// TIA Portal project "Inteligenta_szklarnia" (V15.1)

(* hardware
DEVICE "HMI_test"  KTP700 Basic PN
   slot 0: "HMI_test"  KTP700 Basic PN  6AV2 123-2GB03-0AX0  15.1.0.0
   slot 1: "HMI_RT_1"  KTP700 Basic PN  6AV2 123-2GB03-0AX0  15.1.0.0
   slot 5: "HMI_test.IE_CP_1"  PROFINET Interface  15.0.1.0
      slot 1: "PROFINET Interface_1"  PROFINET Interface
         slot 1: "Port_1"  Port
DEVICE "S7-1200 station_2"  S7-1200 Station
   slot 0: "Rack_0"  S7-1200 Rack  Rack  V1.0
   slot 1: "PLC_1"  CPU 1214C AC/DC/Rly  6ES7 214-1BE30-0XB0  V2.2
DEVICE "HMI_1"  KTP700 Basic PN
   slot 0: "HMI_1"  KTP700 Basic PN  6AV2 123-2GB03-0AX0  15.1.0.0
   slot 1: "HMI_RT_3"  KTP700 Basic PN  6AV2 123-2GB03-0AX0  15.1.0.0
   slot 5: "HMI_1.IE_CP_1"  PROFINET Interface  15.0.1.0
      slot 1: "PROFINET Interface_1"  PROFINET Interface
         slot 1: "Port_1"  Port
DEVICE "S7-1200 station_1"  S7-1200 Station
   slot 0: "Rack_0"  S7-1200 Rack  Rack  V1.0
   slot 1: "PLC_do_symulacji"  CPU 1214C AC/DC/Rly  6ES7 214-1BG40-0XB0  V4.2
DEVICE "HMI_do_symulacji"  KTP700 Basic PN
   slot 0: "HMI_do_symulacji"  KTP700 Basic PN  6AV2 123-2GB03-0AX0  15.1.0.0
   slot 1: "HMI_RT_2"  KTP700 Basic PN  6AV2 123-2GB03-0AX0  15.1.0.0
   slot 5: "HMI_do_symulacji.IE_CP_1"  PROFINET Interface  15.0.1.0
      slot 1: "PROFINET Interface_1"  PROFINET Interface
         slot 1: "Port_1"  Port
*)

// ===== PLC "PLC_1"  CPU 1214C AC/DC/Rly =====

VAR_GLOBAL   // PLC tag table "Default tag table"
   "Tag_1" AT %I0.0 : Bool;
   "Tag_ScreenNumber" AT %MD0 : DInt;
   "FirstScan" AT %M1.0 : Bool;
   "DiagStatusUpdate" AT %M1.1 : Bool;
   "AlwaysTRUE" AT %M1.2 : Bool;
   "AlwaysFALSE" AT %M1.3 : Bool;
END_VAR

VAR_GLOBAL   // PLC tag table "wyjscia"
   "Grzałka" AT %Q0.0 : Bool;
   "Wentylator" AT %Q0.1 : Bool;
   "Pompa_wodna" AT %Q0.2 : Bool;
   "Rolety_zamykanie" AT %Q0.4 : Bool;
   "Alarm_ostrzegwaczy" AT %Q0.5 : Bool;
   "Siłownik_okien_otwieranie" AT %Q0.6 : Bool;
   "Siłownik_okien_zamykanie" AT %Q0.7 : Bool;
   "Rolety_otwieranie" AT %Q0.3 : Bool;
END_VAR

DATA_BLOCK "Parametry"   // DB1
{ S7_Optimized_Access := 'TRUE' }
VERSION : 0.1
   VAR
      Wilgotność_powietrza : Int;
      Wilgotność_gleby : Int;
      temeratura : Real;
      Czujnik_światła : Int;
      Czujnik_wiatru : Int;
      czujnik_CO2 : Int;
      stopien_zasloniecia_rolet : Int;
   END_VAR
BEGIN
END_DATA_BLOCK

DATA_BLOCK "Wejscia_HMI"   // DB2
{ S7_Optimized_Access := 'TRUE' }
VERSION : 0.1
   VAR
      Temperatura : Real;
      CO2 : Real;
      Wilgotność_gleby : Int;
      Wilgotność_powietrza : Int;
      Zaciemnienie : Int;
      naslonecznienie_manual : Int;
   END_VAR
BEGIN
END_DATA_BLOCK

DATA_BLOCK "Receptury"   // DB3
{ S7_Optimized_Access := 'TRUE' }
VERSION : 0.1
   VAR
      nasłonecznienie : Array[0..5] of Int;
      system_okien : Array[0..5] of Bool;
      wilgotnosc_gleby : Array[0..5] of Int;
      wilgotnosc_powietrza : Array[0..5] of Int;
      temperatua : Array[0..5] of Real;
      nazwa : Array[0..5] of String;
   END_VAR
BEGIN
END_DATA_BLOCK

DATA_BLOCK "Archiwizowane_parametry"   // DB4
{ S7_Optimized_Access := 'TRUE' }
VERSION : 0.1
   VAR
      Temperatura : Array[0..335] of Real;
      Wilgotnosc : Array[0..335] of Int;
      Naslonecznienie : Array[0..335] of Int;
      iterator : Int := 0;   // Iterator służący do zapisu danych w odpowiednich komórkach tablicy.
      Zerowanie : Array[0..335] of Int;
   END_VAR
BEGIN
   Naslonecznienie[0] := 0;
   Naslonecznienie[1] := 0;
END_DATA_BLOCK

// folder: System blocks/Program resources

DATA_BLOCK "IEC_Timer_0_DB"   // DB5
{ S7_Optimized_Access := 'TRUE' }
AUTHOR : Simatic
FAMILY : IEC
NAME : IEC_TMR
VERSION : 1.0
// stored: InstanceOfName IEC_TIMER
"IEC_TIMER"
BEGIN
END_DATA_BLOCK

// folder: (top level)

FUNCTION "Rolety" : Void   // FC1, LAD
{ S7_Optimized_Access := 'TRUE' }
VERSION : 0.1
   VAR_INPUT
      Czy_automatyczny : Bool;
      Czy_manualny : Bool;
   END_VAR
   VAR_TEMP   // added for the SCL form of the ladder/FBD networks
      _w1 : Bool;
   END_VAR
BEGIN

REGION Network 1: Sterowanie roletami w trybie automatycznym
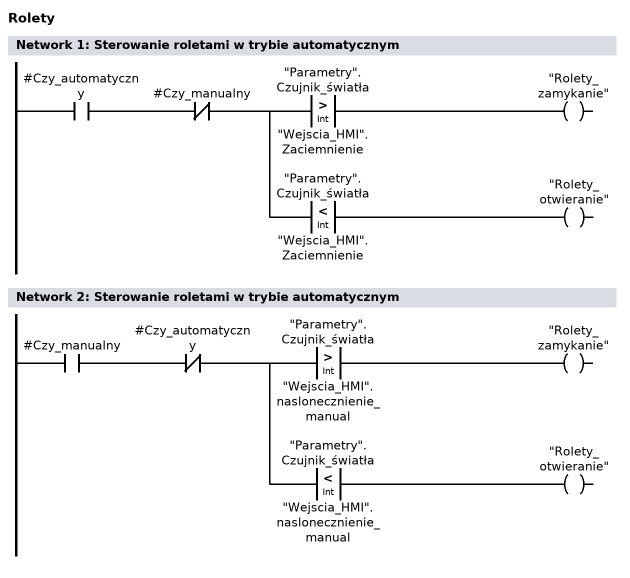
   RUNG wire#powerrail
      Contact( #Czy_automatyczny )
      I_Contact( #Czy_manualny )
      wire#w1
      { S7_Templates := "SrcType := Int" } GT_Contact(in1 := "Parametry".Czujnik_światła, in2 := "Wejscia_HMI".Zaciemnienie)
      Coil( "Rolety_zamykanie" )
   END_RUNG
   RUNG wire#w1
      { S7_Templates := "SrcType := Int" } LT_Contact(in1 := "Parametry".Czujnik_światła, in2 := "Wejscia_HMI".Zaciemnienie)
      Coil( "Rolety_otwieranie" )
   END_RUNG
   // the same network as SCL:
   #_w1 := #Czy_automatyczny AND NOT #Czy_manualny;
   "Rolety_zamykanie" := #_w1 AND ("Parametry".Czujnik_światła > "Wejscia_HMI".Zaciemnienie);
   "Rolety_otwieranie" := #_w1 AND ("Parametry".Czujnik_światła < "Wejscia_HMI".Zaciemnienie);
END_REGION

REGION Network 2: Sterowanie roletami w trybie automatycznym
   RUNG wire#powerrail
      Contact( #Czy_manualny )
      I_Contact( #Czy_automatyczny )
      wire#w1
      { S7_Templates := "SrcType := Int" } GT_Contact(in1 := "Parametry".Czujnik_światła, in2 := "Wejscia_HMI".naslonecznienie_manual)
      Coil( "Rolety_zamykanie" )
   END_RUNG
   RUNG wire#w1
      { S7_Templates := "SrcType := Int" } LT_Contact(in1 := "Parametry".Czujnik_światła, in2 := "Wejscia_HMI".naslonecznienie_manual)
      Coil( "Rolety_otwieranie" )
   END_RUNG
   // the same network as SCL:
   #_w1 := #Czy_manualny AND NOT #Czy_automatyczny;
   "Rolety_zamykanie" := #_w1 AND ("Parametry".Czujnik_światła > "Wejscia_HMI".naslonecznienie_manual);
   "Rolety_otwieranie" := #_w1 AND ("Parametry".Czujnik_światła < "Wejscia_HMI".naslonecznienie_manual);
END_REGION
END_FUNCTION

FUNCTION "Archiwizacja_parametrow" : Void   // FC2, LAD
{ S7_Optimized_Access := 'TRUE' }
VERSION : 0.1
// Zapis parametrów do bloku DB odbywa się co pół godziny. Po uruchomieniu sterownika pierwszy zapis nie odbywa się od razu, aby wykres nie przedstawiał parametrów, które nie były jeszcze regulowane.
BEGIN

REGION Network 1
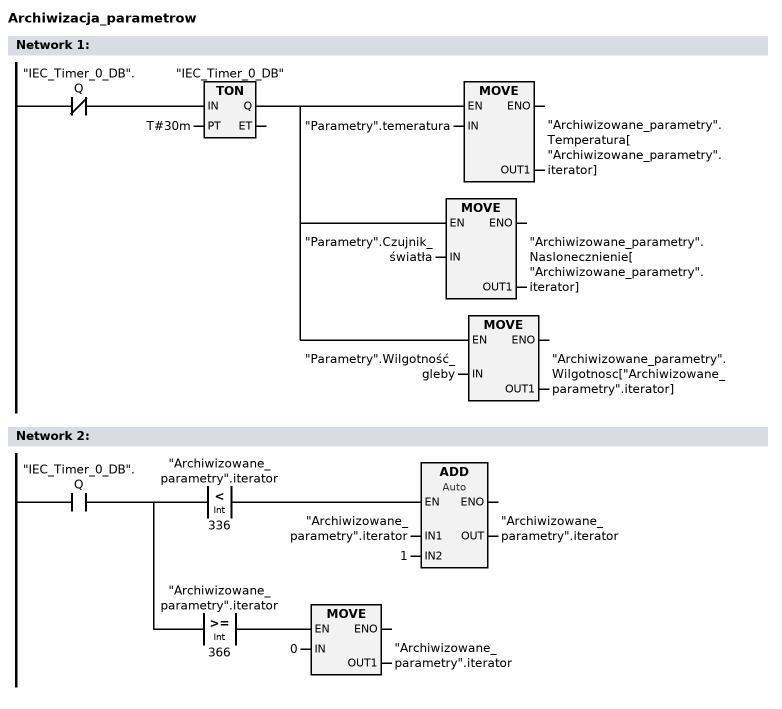
   "IEC_Timer_0_DB".TON(IN := NOT "IEC_Timer_0_DB".Q, PT := T#30m);
   IF "IEC_Timer_0_DB".Q THEN
       "Archiwizowane_parametry".Temperatura["Archiwizowane_parametry".iterator] := "Parametry".temeratura;
       "Archiwizowane_parametry".Naslonecznienie["Archiwizowane_parametry".iterator] := "Parametry".Czujnik_światła;
       "Archiwizowane_parametry".Wilgotnosc["Archiwizowane_parametry".iterator] := "Parametry".Wilgotność_gleby;
   END_IF;
END_REGION

REGION Network 2
   RUNG wire#powerrail
      Contact( "IEC_Timer_0_DB".Q )
      wire#w1
      { S7_Templates := "SrcType := Int" } LT_Contact(in1 := "Archiwizowane_parametry".iterator, in2 := 336)
      { S7_GenerateENO := "TRUE" } Add(in1 := "Archiwizowane_parametry".iterator, in2 := 1, out => "Archiwizowane_parametry".iterator)
   END_RUNG
   RUNG wire#w1
      { S7_Templates := "SrcType := Int" } GE_Contact(in1 := "Archiwizowane_parametry".iterator, in2 := 366)
      { S7_GenerateENO := "TRUE" } Move(in := 0, out1 => "Archiwizowane_parametry".iterator)
   END_RUNG
   // the same network as SCL:
   IF "IEC_Timer_0_DB".Q AND ("Archiwizowane_parametry".iterator < 336) THEN
       "Archiwizowane_parametry".iterator := "Archiwizowane_parametry".iterator + 1;
   END_IF;
   IF "IEC_Timer_0_DB".Q AND ("Archiwizowane_parametry".iterator >= 366) THEN
       "Archiwizowane_parametry".iterator := 0;
   END_IF;
END_REGION
END_FUNCTION

ORGANIZATION_BLOCK "Main"   // OB1, LAD, ProgramCycle
TITLE = "Main Program Sweep (Cycle)"
{ S7_Optimized_Access := 'TRUE' }
VERSION : 0.1
   VAR_INPUT
      Initial_Call : Bool;   // Initial call of this OB
      Remanence : Bool;   // =True, if remanent data are available
   END_VAR
BEGIN

REGION Network 1
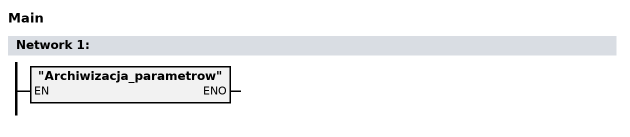
   RUNG wire#powerrail
      "Archiwizacja_parametrow"()
   END_RUNG
   // the same network as SCL:
   "Archiwizacja_parametrow"();
END_REGION
END_ORGANIZATION_BLOCK

ORGANIZATION_BLOCK "Startup"   // OB100, LAD, Startup
TITLE = "Complete Restart"
{ S7_Optimized_Access := 'TRUE' }
VERSION : 0.1
   VAR_INPUT
      LostRetentive : Bool;   // True if retentive data are lost
      LostRTC : Bool;   // True if date and time are lost
   END_VAR
BEGIN

REGION Network 1
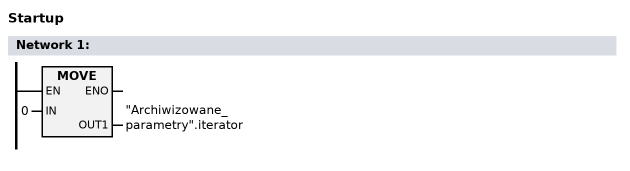
   RUNG wire#powerrail
      { S7_GenerateENO := "TRUE" } Move(in := 0, out1 => "Archiwizowane_parametry".iterator)
   END_RUNG
   // the same network as SCL:
   "Archiwizowane_parametry".iterator := 0;
END_REGION
END_ORGANIZATION_BLOCK

// ===== PLC "PLC_do_symulacji"  CPU 1214C AC/DC/Rly =====

VAR_GLOBAL   // PLC tag table "Default tag table"
   "Tag_1" AT %M0.0 : Bool;
   "System_Byte" AT %MB1 : Byte;
   "FirstScan" AT %M1.0 : Bool;
   "DiagStatusUpdate" AT %M1.1 : Bool;
   "AlwaysTRUE" AT %M1.2 : Bool;
   "AlwaysFALSE" AT %M1.3 : Bool;
   "Tag_2" AT %M0.1 : Bool;
END_VAR

VAR_GLOBAL   // PLC tag table "wyjscia"
   "Grzałka" AT %Q0.0 : Bool;
   "Wentylator" AT %Q0.1 : Bool;
   "Pompa_wodna" AT %Q0.2 : Bool;
   "Rolety_zamykanie" AT %Q0.4 : Bool;
   "Alarm_ostrzegwaczy" AT %Q0.5 : Bool;
   "Siłownik_okien_otwieranie" AT %Q0.6 : Bool;
   "Siłownik_okien_zamykanie" AT %Q0.7 : Bool;
   "Rolety_otwieranie" AT %Q0.3 : Bool;
END_VAR

DATA_BLOCK "Wejscia_PLC"   // DB1
{ S7_Optimized_Access := 'TRUE' }
VERSION : 0.1
   VAR
      Czujnik_wilgotności_powietrza : Int;   // Czujnik wilgotności powietrza w szklarni
      Czujnik_wilgotności_gleby : Int;   // Czujnik wilgotności gleby w szklarni
      Temeratura_wewnetrzna : Real;   // Temperatura wewnątrz szklarni
      Czujnik_natezenia_swiatła : Int;   // Czujnik natężenia światła wewnątrz szklarni
      Czujnik_wiatru : Int;   // Czujnik prędkości wiatru poza szklarnią
      Czujnik_CO2 : Int;   // Czujnik stężenia dwutlenku węgla w szklarni
      Stopien_zasloniecia_rolet : Int;   // Stopień zasłonięcia rolet w szklarni (przyjęty przedział 0-100%)
      Temperatura_zewnetrzna : Int;   // Temperatura mierzona na zewnątrz, poza szklarnią. Typ Int, ponieważ nie jest wymagana taka dokładność jak w pomiarze temperatury wewnętrznej.
   END_VAR
BEGIN
END_DATA_BLOCK

DATA_BLOCK "HMI"   // DB2
{ S7_Optimized_Access := 'TRUE' }
VERSION : 0.1
   VAR
      System_okien_auto : Bool;   // Wł/wył system okien w trybie automatycznym
      Przycisk_pompa_manual : Bool;   // Przycisk pompy w trybie manualnym
      Przycisk_grzanie_manual : Bool;   // Przycisk grzałki w trybie manualnym
      Przycisk_wentylacja_manual : Bool;   // Przycisk wentylacji w trybie manualnym
      Stopien_otwarcia_okien_manual : Int;   // Ustawiony w trybie manualnym stopień otwarcia okien
      Stopien_zasloniecia_rolet_manual : Int;   // Ustawiony w trybie manualnym stopień zasłonięcia rolet
      Temperatura_auto : Real := 22.0;   // Nastawiona temeratura w trybie automatycznym
      Naslonecznienie_auto : Int := 1000;   // Nastawiona wartość nasłonecznienia w trybie automatycznym
      Wilgotnosc_powietrza_auto : Int := 50;   // Nastawiona wartość wilgotności powietrza w trybie automatycznym
      Wilgotnosc_gleby_auto : Int := 60;   // Nastawiona wartość wilgotności gleby w trybie automatycznym
      Przycisk_zatwierdz : Bool;   // Przycisk zatwierdzający wcześniej wybrane ustawienia trybu automatycznego lub receptury
      Numer_ekranu_HMI : Int;   // Numer aktualnie otwartego ekranu w HMI
   END_VAR
BEGIN
END_DATA_BLOCK

DATA_BLOCK "Receptury"   // DB3
{ S7_Optimized_Access := 'TRUE' }
VERSION : 0.1
   VAR
      nasłonecznienie : Array[0..5] of Int;
      system_okien : Array[0..5] of Bool;
      wilgotnosc_gleby : Array[0..5] of Int;
      wilgotnosc_powietrza : Array[0..5] of Int;
      temperatua : Array[0..5] of Real;
      nazwa : Array[0..5] of String;
   END_VAR
BEGIN
END_DATA_BLOCK

DATA_BLOCK "Tryb_auto_parametry"   // DB7
{ S7_Optimized_Access := 'TRUE' }
VERSION : 0.1
   VAR
      Temperatura : Real;
      Naslonecznienie : Int;
      Wilgotnosc_powietrza : Int;
      Wilgotnosc_gleby : Int;
      System_okien : Bool;
   END_VAR
BEGIN
END_DATA_BLOCK

// folder: Archiwizacja_parametrow

DATA_BLOCK "Archiwizowane_parametry"   // DB4
{ S7_Optimized_Access := 'TRUE' }
VERSION : 0.1
   VAR
      Temperatura : Array[0..335] of Real;
      Wilgotnosc : Array[0..335] of Int;
      Naslonecznienie : Array[0..335] of Int;
      iterator : Int := 0;   // Iterator służący do zapisu danych w odpowiednich komórkach tablicy.
   END_VAR
BEGIN
   Naslonecznienie[0] := 0;
   Naslonecznienie[1] := 0;
END_DATA_BLOCK

// folder: System blocks/Program resources

DATA_BLOCK "IEC_Timer_0_DB"   // DB5
{ S7_Optimized_Access := 'TRUE' }
AUTHOR : Simatic
FAMILY : IEC
NAME : IEC_TMR
VERSION : 1.0
// stored: InstanceOfName IEC_TIMER
"IEC_TIMER"
BEGIN
END_DATA_BLOCK

DATA_BLOCK "IEC_Timer_0_DB_1"   // DB6
{ S7_Optimized_Access := 'TRUE' }
AUTHOR : Simatic
FAMILY : IEC
NAME : IEC_TMR
VERSION : 1.0
// stored: InstanceOfName IEC_TIMER
"IEC_TIMER"
BEGIN
END_DATA_BLOCK

// folder: (top level)

FUNCTION "Rolety" : Void   // FC1, LAD
{ S7_Optimized_Access := 'TRUE' }
VERSION : 0.1
   VAR_INPUT
      Czy_automatyczny : Bool;
      Czy_manualny : Bool;
   END_VAR
   VAR_TEMP   // added for the SCL form of the ladder/FBD networks
      _w1 : Bool;
   END_VAR
BEGIN

REGION Network 1: Sterowanie roletami w trybie automatycznym
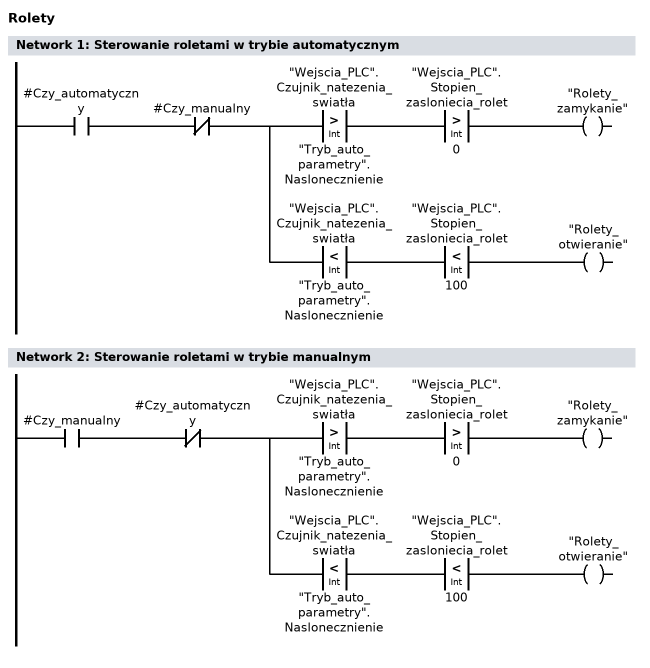
   RUNG wire#powerrail
      Contact( #Czy_automatyczny )
      I_Contact( #Czy_manualny )
      wire#w1
      { S7_Templates := "SrcType := Int" } GT_Contact(in1 := "Wejscia_PLC".Czujnik_natezenia_swiatła, in2 := "Tryb_auto_parametry".Naslonecznienie)
      { S7_Templates := "SrcType := Int" } GT_Contact(in1 := "Wejscia_PLC".Stopien_zasloniecia_rolet, in2 := 0)
      Coil( "Rolety_zamykanie" )
   END_RUNG
   RUNG wire#w1
      { S7_Templates := "SrcType := Int" } LT_Contact(in1 := "Wejscia_PLC".Czujnik_natezenia_swiatła, in2 := "Tryb_auto_parametry".Naslonecznienie)
      { S7_Templates := "SrcType := Int" } LT_Contact(in1 := "Wejscia_PLC".Stopien_zasloniecia_rolet, in2 := 100)
      Coil( "Rolety_otwieranie" )
   END_RUNG
   // the same network as SCL:
   #_w1 := #Czy_automatyczny AND NOT #Czy_manualny;
   "Rolety_zamykanie" := #_w1 AND ("Wejscia_PLC".Czujnik_natezenia_swiatła > "Tryb_auto_parametry".Naslonecznienie) AND ("Wejscia_PLC".Stopien_zasloniecia_rolet > 0);
   "Rolety_otwieranie" := #_w1 AND ("Wejscia_PLC".Czujnik_natezenia_swiatła < "Tryb_auto_parametry".Naslonecznienie) AND ("Wejscia_PLC".Stopien_zasloniecia_rolet < 100);
END_REGION

REGION Network 2: Sterowanie roletami w trybie manualnym
   RUNG wire#powerrail
      Contact( #Czy_manualny )
      I_Contact( #Czy_automatyczny )
      wire#w1
      { S7_Templates := "SrcType := Int" } GT_Contact(in1 := "Wejscia_PLC".Czujnik_natezenia_swiatła, in2 := "Tryb_auto_parametry".Naslonecznienie)
      { S7_Templates := "SrcType := Int" } GT_Contact(in1 := "Wejscia_PLC".Stopien_zasloniecia_rolet, in2 := 0)
      Coil( "Rolety_zamykanie" )
   END_RUNG
   RUNG wire#w1
      { S7_Templates := "SrcType := Int" } LT_Contact(in1 := "Wejscia_PLC".Czujnik_natezenia_swiatła, in2 := "Tryb_auto_parametry".Naslonecznienie)
      { S7_Templates := "SrcType := Int" } LT_Contact(in1 := "Wejscia_PLC".Stopien_zasloniecia_rolet, in2 := 100)
      Coil( "Rolety_otwieranie" )
   END_RUNG
   // the same network as SCL:
   #_w1 := #Czy_manualny AND NOT #Czy_automatyczny;
   "Rolety_zamykanie" := #_w1 AND ("Wejscia_PLC".Czujnik_natezenia_swiatła > "Tryb_auto_parametry".Naslonecznienie) AND ("Wejscia_PLC".Stopien_zasloniecia_rolet > 0);
   "Rolety_otwieranie" := #_w1 AND ("Wejscia_PLC".Czujnik_natezenia_swiatła < "Tryb_auto_parametry".Naslonecznienie) AND ("Wejscia_PLC".Stopien_zasloniecia_rolet < 100);
END_REGION
END_FUNCTION

FUNCTION "TO_DO_Sterowanie_temperatura" : Void   // FC3, LAD
{ S7_Optimized_Access := 'TRUE' }
VERSION : 0.1
   VAR_INPUT
      czy_manualny : Bool;
      czy_automatyczny : Bool;
   END_VAR
   VAR_TEMP
      Histereza_minus : Real;   // Wartość zadanej temperatury zmieniona o dolną wartość hiterezy
      Histereza_plus : Real;   // Wartość zadanej temperatury zmieniona o górną wartość hiterezy
   END_VAR
   VAR_TEMP   // added for the SCL form of the ladder/FBD networks
      _w1 : Bool;
   END_VAR
BEGIN

REGION Network 1: Sterowanie temperaturą w trybie automatycznym
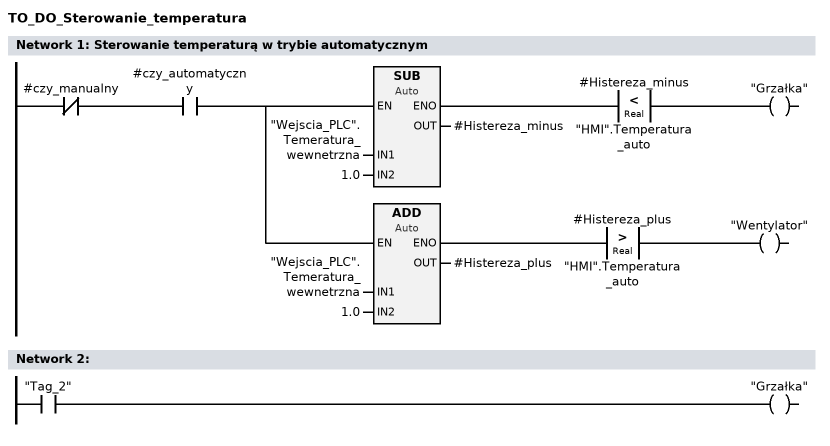
   RUNG wire#powerrail
      I_Contact( #czy_manualny )
      Contact( #czy_automatyczny )
      wire#w1
      Sub(in1 := "Wejscia_PLC".Temeratura_wewnetrzna, in2 := 1.0, out => #Histereza_minus)
      { S7_Templates := "SrcType := Real" } LT_Contact(in1 := #Histereza_minus, in2 := "HMI".Temperatura_auto)
      Coil( "Grzałka" )
   END_RUNG
   RUNG wire#w1
      Add(in1 := "Wejscia_PLC".Temeratura_wewnetrzna, in2 := 1.0, out => #Histereza_plus)
      { S7_Templates := "SrcType := Real" } GT_Contact(in1 := #Histereza_plus, in2 := "HMI".Temperatura_auto)
      Coil( "Wentylator" )
   END_RUNG
   // the same network as SCL:
   #_w1 := NOT #czy_manualny AND #czy_automatyczny;
   IF #_w1 THEN #Histereza_minus := "Wejscia_PLC".Temeratura_wewnetrzna - 1.0; END_IF;
   "Grzałka" := #_w1 AND (#Histereza_minus < "HMI".Temperatura_auto);
   IF #_w1 THEN #Histereza_plus := "Wejscia_PLC".Temeratura_wewnetrzna + 1.0; END_IF;
   "Wentylator" := #_w1 AND (#Histereza_plus > "HMI".Temperatura_auto);
END_REGION

REGION Network 2
   RUNG wire#powerrail
      Contact( "Tag_2" )
      Coil( "Grzałka" )
   END_RUNG
   // the same network as SCL:
   "Grzałka" := "Tag_2";
END_REGION
END_FUNCTION

FUNCTION "Zapis_parametrow_trybu_auto" : Void   // FC4, LAD
{ S7_Optimized_Access := 'TRUE' }
VERSION : 0.1
   VAR_TEMP   // added for the SCL form of the ladder/FBD networks
      _w1 : Bool;
   END_VAR
BEGIN

REGION Network 1: Zapis wybranych na HMI parametrów, aby zostały one stałe do kolejnego zatwierdzenia ich zmiany.
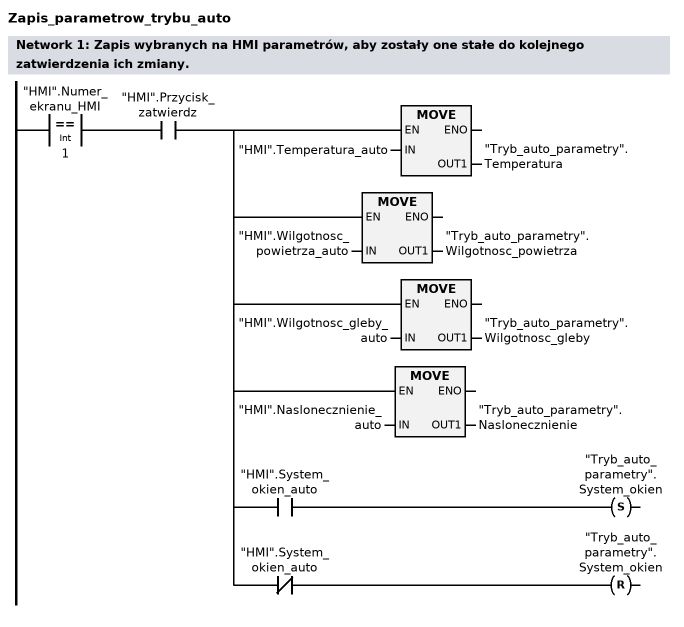
   RUNG wire#powerrail
      { S7_Templates := "SrcType := Int" } EQ_Contact(in1 := "HMI".Numer_ekranu_HMI, in2 := 1)
      Contact( "HMI".Przycisk_zatwierdz )
      wire#w1
      Move(in := "HMI".Temperatura_auto, out1 => "Tryb_auto_parametry".Temperatura)
   END_RUNG
   RUNG wire#w1
      Move(in := "HMI".Wilgotnosc_powietrza_auto, out1 => "Tryb_auto_parametry".Wilgotnosc_powietrza)
   END_RUNG
   RUNG wire#w1
      Move(in := "HMI".Wilgotnosc_gleby_auto, out1 => "Tryb_auto_parametry".Wilgotnosc_gleby)
   END_RUNG
   RUNG wire#w1
      Move(in := "HMI".Naslonecznienie_auto, out1 => "Tryb_auto_parametry".Naslonecznienie)
   END_RUNG
   RUNG wire#w1
      Contact( "HMI".System_okien_auto )
      S_Coil( "Tryb_auto_parametry".System_okien )
   END_RUNG
   RUNG wire#w1
      I_Contact( "HMI".System_okien_auto )
      R_Coil( "Tryb_auto_parametry".System_okien )
   END_RUNG
   // the same network as SCL:
   #_w1 := ("HMI".Numer_ekranu_HMI = 1) AND "HMI".Przycisk_zatwierdz;
   IF #_w1 THEN
       "Tryb_auto_parametry".Temperatura := "HMI".Temperatura_auto;
       "Tryb_auto_parametry".Wilgotnosc_powietrza := "HMI".Wilgotnosc_powietrza_auto;
       "Tryb_auto_parametry".Wilgotnosc_gleby := "HMI".Wilgotnosc_gleby_auto;
       "Tryb_auto_parametry".Naslonecznienie := "HMI".Naslonecznienie_auto;
   END_IF;
   IF #_w1 AND "HMI".System_okien_auto THEN "Tryb_auto_parametry".System_okien := TRUE; END_IF;
   IF #_w1 AND NOT "HMI".System_okien_auto THEN "Tryb_auto_parametry".System_okien := FALSE; END_IF;
END_REGION
END_FUNCTION

ORGANIZATION_BLOCK "Main"   // OB1, LAD, ProgramCycle
TITLE = "Main Program Sweep (Cycle)"
{ S7_Optimized_Access := 'TRUE' }
VERSION : 0.1
   VAR_INPUT
      Initial_Call : Bool;   // Initial call of this OB
      Remanence : Bool;   // =True, if remanent data are available
   END_VAR
BEGIN

REGION Network 1
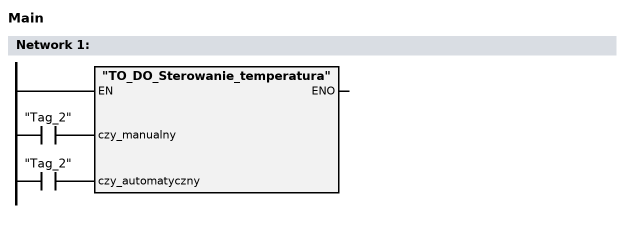
   RUNG wire#powerrail
      "TO_DO_Sterowanie_temperatura"(czy_manualny := wire#w1, czy_automatyczny := wire#w2)
   END_RUNG
   RUNG wire#powerrail
      Contact( "Tag_2" )
   END_RUNG wire#w1
   RUNG wire#powerrail
      Contact( "Tag_2" )
   END_RUNG wire#w2
   // the same network as SCL:
   "TO_DO_Sterowanie_temperatura"(czy_manualny := "Tag_2", czy_automatyczny := "Tag_2");
END_REGION
END_ORGANIZATION_BLOCK

// folder: Archiwizacja_parametrow

FUNCTION "Archiwizacja_parametrow" : Void   // FC2, LAD
{ S7_Optimized_Access := 'TRUE' }
VERSION : 0.1
// Zapis parametrów do bloku DB odbywa się co pół godziny. Po uruchomieniu sterownika pierwszy zapis nie odbywa się od razu, aby wykres nie przedstawiał parametrów, które nie były jeszcze regulowane. Oczytane watosci zapisywane są w tablicach w bloku DB.
   VAR CONSTANT
      iterator : Int := 0;
   END_VAR
   VAR_TEMP   // added for the SCL form of the ladder/FBD networks
      _w1 : Bool;
   END_VAR
BEGIN

REGION Network 1
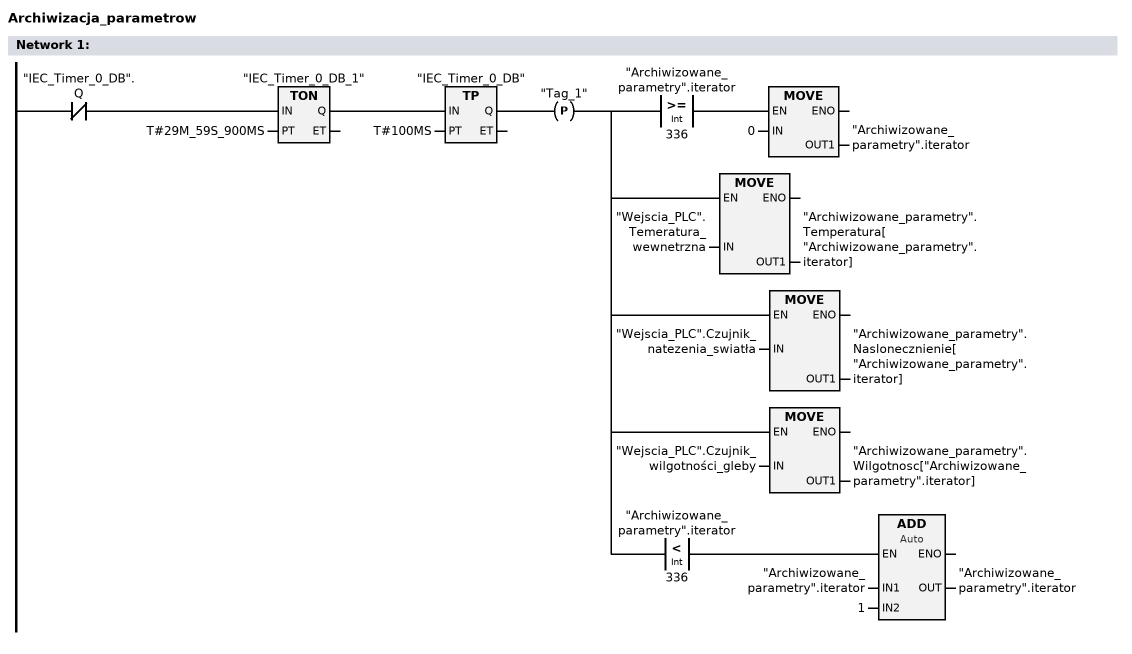
   "IEC_Timer_0_DB_1".TON(IN := NOT "IEC_Timer_0_DB".Q, PT := T#29M_59S_900MS);
   "IEC_Timer_0_DB".TP(IN := "IEC_Timer_0_DB_1".Q, PT := T#100MS);
   #_w1 := "IEC_Timer_0_DB".Q AND NOT "Tag_1";   // rising edge
   "Tag_1" := "IEC_Timer_0_DB".Q;
   IF #_w1 AND ("Archiwizowane_parametry".iterator >= 336) THEN
       "Archiwizowane_parametry".iterator := 0;
   END_IF;
   IF #_w1 THEN
       "Archiwizowane_parametry".Temperatura["Archiwizowane_parametry".iterator] := "Wejscia_PLC".Temeratura_wewnetrzna;
       "Archiwizowane_parametry".Naslonecznienie["Archiwizowane_parametry".iterator] := "Wejscia_PLC".Czujnik_natezenia_swiatła;
       "Archiwizowane_parametry".Wilgotnosc["Archiwizowane_parametry".iterator] := "Wejscia_PLC".Czujnik_wilgotności_gleby;
   END_IF;
   IF #_w1 AND ("Archiwizowane_parametry".iterator < 336) THEN
       "Archiwizowane_parametry".iterator := "Archiwizowane_parametry".iterator + 1;
   END_IF;
END_REGION
END_FUNCTION

(* ===== HMI "HMI_RT_1" =====
system functions are stored by id; their names below are inferred from use
connection "HMI_Connection_2": 
connection "HMI_Connection_1": 
connection "Connection_1": ETHERNET, SMART_S7_1200_OMS

HMI tags "wyjsciaPLC"
   "Alarm_ostrzegwaczy" : Bool = PLC Alarm_ostrzegwaczy AT %Q0.5, 100 ms
   "Grzałka" : Bool = PLC Grzałka AT %Q0.0, 100 ms
   "Pompa_wodna" : Bool = PLC Pompa_wodna AT %Q0.2, 100 ms
   "Rolety_otwieranie" : Bool = PLC Rolety_otwieranie AT %Q0.3, 100 ms
   "Rolety_zamykanie" : Bool = PLC Rolety_zamykanie AT %Q0.4, 100 ms
   "Siłownik_okien_otwieranie" : Bool = PLC Siłownik_okien_otwieranie AT %Q0.6, 100 ms
   "Siłownik_okien_zamykanie" : Bool = PLC Siłownik_okien_zamykanie AT %Q0.7, 100 ms
   "Wentylator" : Bool = PLC Wentylator AT %Q0.1, 100 ms
   "Tag_ScreenNumber" : DInt = PLC Tag_ScreenNumber AT %MD0, 500 ms
   "Parametry_Czujnik_światła" : Int = PLC Parametry.Czujnik_światła, 500 ms
   "Parametry_temeratura" : Real = PLC Parametry.temeratura, 500 ms
   "Parametry_Czujnik_wiatru" : Int = PLC Parametry.Czujnik_wiatru, 500 ms
   "Parametry_Wilgotność_powietrza" : Int = PLC Parametry.Wilgotność_powietrza, 500 ms
   "Parametry_czujnik_CO2" : Int = PLC Parametry.czujnik_CO2, 500 ms
   "Parametry_Wilgotność_gleby" : Int = PLC Parametry.Wilgotność_gleby, 500 ms
   "Wejscia_HMI_Temperatura" : Real = PLC Wejscia_HMI.Temperatura, 500 ms
   "Parametry_stopien_zasloniecia_rolet" : Int = PLC Parametry.stopien_zasloniecia_rolet, 1 s
   "Wejscia_HMI_Zaciemnienie" : Int = PLC Wejscia_HMI.Zaciemnienie, 1 s
   "Receptury_nazwa{0}" : String[254] = PLC Receptury.nazwa[0], 1 s
   "Receptury_nazwa{1}" : String[254] = PLC Receptury.nazwa[1], 1 s
   "Receptury_nazwa{2}" : String[254] = PLC Receptury.nazwa[2], 1 s
   "Receptury_nazwa{3}" : String[254] = PLC Receptury.nazwa[3], 1 s
   "Receptury_nazwa{4}" : String[254] = PLC Receptury.nazwa[4], 1 s
   "Receptury_nazwa{5}" : String[254] = PLC Receptury.nazwa[5], 1 s

HMI tags "USTAWIENIA_HMI"
   "temperatura_ustawiona_man" : Real, internal
   "stopien_otwarcia_okien_man" : Real, internal
   "wilgotnosc_powietrza_man" : Real, internal
   "wilgotnosc_gleby_man" : Real, internal
   "naslonecznienie_man" : Real, internal
   "nazwa_receptury" : WString[10], internal
   "system_okien" : Bool, internal
   "AlwaysTRUE" : Bool = PLC AlwaysTRUE AT %M1.2, 1 s

Template "Template_1" 800x480
   Button "Exit" at 671,429 size 71x50; TextOff 'Exit'; PictureOff "ExitRuntime_KTP700_Basic_PN_TR"; PictureOn "ExitRuntime_KTP700_Basic_PN_TR"
      on Release: StopRuntime(0)
   Button "Alarms" at 524,429 size 71x50; TextOff 'Alarms'; PictureOff "AlarmDisplay_KTP700_Basic_PN_TR"; PictureOn "AlarmDisplay_KTP700_Basic_PN_TR"
      on Release: function_ef3f5d25("Alarm window_Unacknowledged", -1)
   Button "Start screen" at 169,429 size 71x50; TextOff 'Start screen'; PictureOff "NavigateHome_KTP700_Basic_PN_TR"; PictureOn "NavigateHome_KTP700_Basic_PN_TR"
      on Release: ActivateScreen("Root screen", 0)
      Visibility <- "AlwaysTRUE"
   Button "Language" at 377,429 size 71x50; TextOn 'Language'; TextOff 'Language'; PictureOn "ToggleLanguage_KTP700_Basic_PN_TR"; PictureOff "ToggleLanguage_KTP700_Basic_PN_TR"
      on Release: function_fb9197e8(-1)

screen "Root screen" 800x480, template "Template_1"
   on GenerateScreen: SetTag("Tag_ScreenNumber", 1)
   Button "Button_3" at 10,270 size 300x90; TextOff 'ZAPISZ NOWĄ RECEPTURĘ'
      on Click: ActivateScreen("zapisz_recepture", 0)
   Button "Button_1" at 10,170 size 300x90; TextOff 'TRYB MANUALNY'
      on Click: ActivateScreen("tryb_manualny", 0)
   Button "Button_2" at 10,70 size 301x90; TextOff 'TRYB AUTOMATYCZNY'
      on Click: ActivateScreen("tryb_automatyczny", 0)
   TextField "Text field_2" at 32,2 size 738x63; Text 'AUTOMATYCZNA SZKLARNIA'
   GraphicView "Graphic view_1" at 370,70 size 392x338; Picture "garden-tools-graphic-clipart-design-free-png"
   Button "Button_4" at 10,370 size 301x90; TextOff 'WYBIERZ RECEPTURĘ'
      on Click: ActivateScreen("wybierz_recepture", 0)
   TextField "Text field_1" at 117,454 size 235x26; Text 'Tego przycisku w symulacji nie widac ale nie chciałem uswac jakby jednak był potrzebny xd'
      Visibility <- "AlwaysTRUE"

screen "zapisz_recepture" 800x480
   TextField "Text field_1" at 282,4 size 253x34; Text 'ZAPISZ RECEPTURE / ZAPISZ RECEPTURĘ'
   Button "Button_1" at 750,0 size 50x50; TextOff 'WRÓĆ'; PictureOff "Back_arrow"
      on Click: function_efd93a16()
   Button "Button_2" at 406,414 size 371x53; TextOff 'ZATWIERDŹ'
      on Click: ActivateScreen("praca", 0)
   Bar "Bar_1" at 17,122 size 70x314; MinimumValue 0; MaximumValue 45
      ProcessValue <- "temperatura_ustawiona_man"
   TextField "Text field_2" at 30,64 size 132x23; Text 'TEMPERATURA'
   Bar "Bar_2" at 223,133 size 54x113; MinimumValue 0; MaximumValue 100
      ProcessValue <- "wilgotnosc_powietrza_man"
   TextField "Text field_3" at 231,45 size 122x42; Text 'WOLGOTNOŚĆ POWIETRZA'
   Button "Button_3" at 115,140 size 73x45; TextOff '+ / +0.5 °C'
      on Press: function_dd21b452("temperatura_ustawiona_man", 0.5)
   Button "Button_7" at 115,201 size 73x45; TextOff '- / -0.5 °C'
      on Press: function_b9b71300("temperatura_ustawiona_man", 0.5)
   TextField "Text field_8" at 93,325 size 109x42; Text 'ustawiona wartość USTAWIONA'
   IOField "I/O field_2" at 106,365 size 62x40; FormatPattern 99.9
      ProcessValue <- "temperatura_ustawiona_man"
   TextField "Text field_11" at 156,367 size 37x37; Text '°C'
   Bar "Bar_4" at 225,346 size 57x127; MinimumValue 0; MaximumValue 100
      ProcessValue <- "wilgotnosc_gleby_man"
   TextField "Text field_10" at 229,254 size 122x42; Text 'WOLGOTNOŚĆ GLEBY'
   Button "Button_8" at 230,300 size 40x40; TextOff '+'
      on Click: function_dd21b452("wilgotnosc_gleby_man", 2)
   Button "Button_9" at 318,300 size 40x40; TextOff '-'
      on Click: function_b9b71300("wilgotnosc_gleby_man", 2)
   IOField "I/O field_5" at 291,401 size 62x40; FormatPattern 999
      ProcessValue <- "wilgotnosc_gleby_man"
   TextField "Text field_12" at 285,384 size 83x20; Text 'USTAWIONA'
   TextField "Text field_14" at 338,404 size 30x29; Text '%'
   Button "Button_10" at 223,87 size 40x40; TextOff '+'
      on Click: function_dd21b452("wilgotnosc_powietrza_man", 5)
   Button "Button_11" at 311,87 size 40x40; TextOff '-'
      on Click: function_b9b71300("wilgotnosc_powietrza_man", 5)
   IOField "I/O field_4" at 291,180 size 62x40; FormatPattern 999
      ProcessValue <- "wilgotnosc_powietrza_man"
   TextField "Text field_16" at 288,167 size 83x20; Text 'USTAWIONA'
   TextField "Text field_18" at 342,184 size 30x29; Text '%'
   Button "Button_14" at 3,1 size 43x43; TextOff 'DOM'; PictureOff "home_1"
      on Click: ActivateScreen("Root screen", 0)
   TextField "Text field_4" at 529,47 size 128x23; Text 'SYSTEM OKIEN'
   Switch "Switch_1" at 503,78 size 185x35; CaptionText 'Switch'; TextOff 'OFF'; TextOn 'ON'
      ProcessValue <- "system_okien"
   IOField "I/O field_1" at 426,311 size 328x81; FormatPattern ????????????????????
      ProcessValue <- "nazwa_receptury"
   TextField "Text field_7" at 406,273 size 380x37; Text 'WPISZ NAZWĘ RECEPTURY'
   GraphicView "Graphic view_1" at 385,338 size 36x30; Picture "Graphic_4"
   GraphicView "Graphic view_2" at 753,338 size 36x30; Picture "Graphic_5"
   TextField "Text field_9" at 387,146 size 161x61; Text 'STOPIEŃ OTWARCIA OKIEN ŚREDNIE NASŁONECZNIENIE'
   Bar "Bar_6" at 404,213 size 373x52; MinimumValue 0; MaximumValue 1500
      ProcessValue <- "naslonecznienie_man"
   Button "Button_4" at 697,145 size 80x50; TextOff '+ / -'
      on Click: function_b9b71300("naslonecznienie_man", 5)
   Button "Button_5" at 589,145 size 80x50; TextOff '- / +'
      on Press: function_dd21b452("naslonecznienie_man", 5)

screen "tryb_manualny" 800x480
   Button "Button_2" at 355,415 size 431x53; TextOff 'ZATWIERDŹ'
      on Click: ActivateScreen("praca", 0)
   TextField "Text field_1" at 282,4 size 223x34; Text 'TRYB MANUALNY'
   Bar "Bar_1" at 181,300 size 60x172; MinimumValue 0; MaximumValue 45
      ProcessValue <- "Parametry_temeratura"
   TextField "Text field_2" at 188,267 size 132x23; Text 'TEMPERATURA'
   Bar "Bar_2" at 181,93 size 60x160; MinimumValue 0; MaximumValue 100
      ProcessValue <- "Parametry_Wilgotność_powietrza"
   TextField "Text field_3" at 198,45 size 122x42; Text 'WOLGOTNOŚĆ POWIETRZA WILGOTNOŚĆ POWIETRZA'
   Bar "Bar_3" at 576,166 size 170x52; MinimumValue 0
      ProcessValue <- "stopien_otwarcia_okien_man"
   TextField "Text field_4" at 576,43 size 186x61; Text 'STOPIEŃ OTWARCIA OKIEN STOPIEŃ OTWARCIA OKIEN'
   IOField "I/O field_1" at 244,368 size 95x40; FormatPattern 99.9
      ProcessValue <- "Wejscia_HMI_Temperatura"
   Bar "Bar_4" at 8,93 size 60x160; MinimumValue 0; MaximumValue 100
      ProcessValue <- "Parametry_Wilgotność_gleby"
   Button "Button_4" at 406,253 size 80x60; TextOff 'PODLEWANIE'
      on Click: InvertBit("Pompa_wodna")
   Button "Button_5" at 536,253 size 80x60; TextOff 'GRZANIE'
      on Click: InvertBit("Grzałka")
   Button "Button_6" at 666,253 size 80x60; TextOff 'WENTYLACJA'
      on Click: InvertBit("Wentylator")
   GraphicView "Graphic view_1" at 675,320 size 60x60; Picture "fan_4829316"
      Visibility <- "Wentylator"
   GraphicView "Graphic view_6" at 545,320 size 60x60; Picture "heater_4463010"
      Visibility <- "Grzałka"
   GraphicView "Graphic view_7" at 415,320 size 60x60; Picture "irrigation_18631825"
      Visibility <- "Pompa_wodna"
   GraphicView "Graphic view_9" at 676,320 size 60x60; Picture "fan_off"
      Visibility <- "Wentylator"
   GraphicView "Graphic view_10" at 546,320 size 60x60; Picture "heater_off"
      Visibility <- "Grzałka"
   GraphicView "Graphic view_11" at 415,320 size 60x60; Picture "irrigation_off"
      Visibility <- "Pompa_wodna"
   TextField "Text field_10" at 18,45 size 122x42; Text 'WOLGOTNOŚĆ GLEBY WILGOTNOŚĆ GLEBY'
   IOField "I/O field_3" at 760,171 size 33x36; FormatPattern 9
      ProcessValue <- "stopien_otwarcia_okien_man"
   IOField "I/O field_6" at 70,148 size 62x40; FormatPattern 999
      ProcessValue <- "Parametry_Wilgotność_gleby"
   TextField "Text field_15" at 115,152 size 35x34; Text '%'
   IOField "I/O field_7" at 252,151 size 62x40; FormatPattern 999
      ProcessValue <- "Parametry_Wilgotność_powietrza"
   TextField "Text field_19" at 294,154 size 35x34; Text '%'
   Button "Button_12" at 576,99 size 50x50; TextOff '+'
      on Click: function_dd21b452("stopien_otwarcia_okien_man", 1)
   Button "Button_13" at 696,98 size 50x50; TextOff '-'
      on Click: function_b9b71300("stopien_otwarcia_okien_man", 1)
   Button "Button_14" at 3,1 size 43x43; TextOff 'DOM'; PictureOff "home_1"
      on Click: ActivateScreen("Root screen", 0)
   Button "Button_1" at 750,0 size 50x50; TextOff 'Text'; PictureOff "Back_arrow"
      on Click: function_efd93a16()
   TextField "Text field_9" at 293,369 size 35x34; Text '°C'
   Circle "Circle_1" at 386,336 size 25x25
      Visibility <- "Pompa_wodna"
   Circle "Circle_4" at 386,336 size 25x25
      Visibility <- "Pompa_wodna"
   Circle "Circle_2" at 511,336 size 25x25
      Visibility <- "Grzałka"
   Circle "Circle_5" at 511,336 size 25x25
      Visibility <- "Grzałka"
   Circle "Circle_3" at 639,336 size 25x25
      Visibility <- "Wentylator"
   Circle "Circle_6" at 639,336 size 25x25
      Visibility <- "Wentylator"
   Bar "Bar_5" at 10,300 size 60x172; MinimumValue 0; MaximumValue 1500
      ProcessValue <- "Parametry_Czujnik_światła"
   TextField "Text field_5" at 3,268 size 161x23; Text 'TEMPERATURA / NASŁONECZNIENIE'
   IOField "I/O field_2" at 70,368 size 95x40; FormatPattern 9999
      ProcessValue <- "Parametry_Czujnik_światła"
   TextField "Text field_6" at 127,356 size 35x64; Text '°C W m'
   TextField "Text field_7" at 152,391 size 31x17; Text '2'
   TextField "Text field_8" at 348,43 size 206x61; Text 'STOPIEŃ OTWARCIA OKIEN STOPIEŃ ZASŁONIENIA ROLET'
   Bar "Bar_6" at 366,166 size 170x52; MinimumValue 0; MaximumValue 100
      ProcessValue <- "naslonecznienie_man"
   Button "Button_3" at 456,98 size 80x50; TextOff '+ / ODSŁOŃ'
      on Click: function_b9b71300("naslonecznienie_man", 5)
   Button "Button_7" at 366,98 size 80x50; TextOff '- / ZASŁOŃ'
      on Press: function_dd21b452("naslonecznienie_man", 5)

screen "wybierz_recepture" 800x480
   TextField "Text field_2" at 257,4 size 280x34; Text 'WYBIERZ RECEPTURE / WYBIERZ RECEPTURĘ'
   Button "Button_1" at 750,0 size 50x50; TextOff 'WRÓĆ'; PictureOff "Back_arrow"
      on Click: function_efd93a16()
   Button "Button_14" at 3,1 size 43x43; TextOff 'DOM'; PictureOff "home_1"
      on Click: ActivateScreen("Root screen", 0)
   TextField "Text field_1" at 18,52 size 23x39; Text '1'
   TextField "Text field_3" at 18,108 size 23x39; Text '2'
   TextField "Text field_4" at 18,169 size 23x39; Text '3'
   TextField "Text field_5" at 18,231 size 23x39; Text '4'
   TextField "Text field_6" at 18,290 size 23x39; Text '5'
   TextField "Text field_7" at 18,351 size 23x39; Text '6'
   Button "Button_2" at 13,415 size 775x55; TextOff '-ZATWIERDŹ-'
      on Click: ActivateScreen("praca", 0)
   Button "Button_3" at 720,68 size 60x60; TextOff 'Text'; PictureOff "Double_up_arrow"
   Button "Button_4" at 720,162 size 60x60; TextOff 'Text'; PictureOff "Double_down_arrow"
   Button "Button_5" at 708,326 size 83x64; TextOff 'USUŃ'
   IOField "I/O field_1" at 90,58 size 243x32; FormatPattern ????????????????????
      ProcessValue <- "Receptury_nazwa{0}"
   IOField "I/O field_2" at 90,115 size 241x32; FormatPattern ????????????????????
      ProcessValue <- "Receptury_nazwa{1}"
   IOField "I/O field_3" at 90,176 size 267x32; FormatPattern ????????????????????
      ProcessValue <- "Receptury_nazwa{2}"
   IOField "I/O field_4" at 90,238 size 264x32; FormatPattern ????????????????????
      ProcessValue <- "Receptury_nazwa{3}"
   IOField "I/O field_5" at 90,294 size 230x32; FormatPattern ????????????????????
      ProcessValue <- "Receptury_nazwa{4}"
   IOField "I/O field_6" at 90,358 size 506x32; FormatPattern ????????????????????
      ProcessValue <- "Receptury_nazwa{5}"

screen "praca" 800x480
   GraphicView "Graphic view_2" at 28,217 size 100x100; Picture "Thermometer_icon"
   GraphicView "Graphic view_4" at 276,362 size 100x100; Picture "soil-sensor_11298794"
   GraphicView "Graphic view_3" at 28,74 size 100x100; Picture "sensor_4212513"
   GraphicView "Graphic view_5" at 276,75 size 100x100; Picture "sensor_4212519"
   GraphicView "Graphic view_1" at 559,362 size 100x100; Picture "fan_4829316"
      Visibility <- "Wentylator"
   GraphicView "Graphic view_6" at 560,217 size 100x100; Picture "heater_4463010"
      Visibility <- "Grzałka"
   GraphicView "Graphic view_7" at 560,75 size 100x100; Picture "irrigation_18631825"
      Visibility <- "Pompa_wodna"
   GraphicView "Graphic view_8" at 28,362 size 100x100; Picture "anemometer_1113716"
   GraphicView "Graphic view_9" at 560,362 size 100x100; Picture "fan_off"
      Visibility <- "Wentylator"
   GraphicView "Graphic view_10" at 561,217 size 100x100; Picture "heater_off"
      Visibility <- "Grzałka"
   GraphicView "Graphic view_11" at 561,75 size 100x100; Picture "irrigation_off"
      Visibility <- "Pompa_wodna"
   GraphicView "Graphic view_12" at 276,217 size 100x100; Picture "sensor_2828470"
   TextField "Text field_1" at 54,52 size 204x23; Text 'INSOLATION / NASŁONECZNIENIE / SONNENEINSTRAHLUNG'
   TextField "Text field_2" at 67,194 size 132x23; Text 'TEMPERATURA'
   TextField "Text field_3" at 46,334 size 166x23; Text 'SZYBKOŚĆ WIATRU'
   TextField "Text field_4" at 349,194 size 123x23; Text 'STĘŻENIE CO2'
   TextField "Text field_5" at 294,50 size 223x23; Text 'WILGOTNOŚĆ POWIETRZA'
   TextField "Text field_6" at 321,339 size 175x23; Text 'WILGOTNOŚĆ GLEBY'
   TextField "Text field_7" at 626,46 size 116x23; Text 'PODLEWANIE'
   TextField "Text field_8" at 643,192 size 80x23; Text 'GRZANIE'
   TextField "Text field_9" at 626,330 size 117x23; Text 'WENTYLACJA'
   TextField "Text field_10" at 282,4 size 256x34; Text 'PODGLĄD NA ŻYWO'
   Button "Button_1" at 750,0 size 50x50; TextOff 'WRÓĆ'; PictureOff "Back_arrow"
      on Click: function_efd93a16()
   Button "Button_2" at 3,1 size 43x43; TextOff 'DOM'; PictureOff "home_1"
      on Click: ActivateScreen("Root screen", 0)
   IOField "I/O field_2" at 120,233 size 97x65; FormatPattern 99.99
      ProcessValue <- "Parametry_temeratura"
   IOField "I/O field_3" at 136,383 size 70x65; FormatPattern 999
      ProcessValue <- "Parametry_Czujnik_wiatru"
   IOField "I/O field_5" at 377,235 size 83x65; FormatPattern 9999
      ProcessValue <- "Parametry_czujnik_CO2"
   TextField "Text field_11" at 214,241 size 46x46; Text '°C'
   IOField "I/O field_4" at 406,95 size 69x65; FormatPattern 999
      ProcessValue <- "Parametry_Wilgotność_powietrza"
   IOField "I/O field_6" at 406,384 size 68x65; FormatPattern 999
      ProcessValue <- "Parametry_Wilgotność_gleby"
   TextField "Text field_12" at 472,106 size 47x46; Text '%'
   TextField "Text field_13" at 472,396 size 47x46; Text '%'
   TextField "Text field_14" at 219,90 size 47x72; Text 'W m²'
   IOField "I/O field_1" at 119,109 size 101x32; FormatPattern 99999
      ProcessValue <- "Parametry_Czujnik_światła"
   TextField "Text field_15" at 210,376 size 52x72; Text 'Km h'
   Circle "Circle_1" at 695,101 size 48x48
      Visibility <- "Pompa_wodna"
   Circle "Circle_2" at 695,243 size 48x48
      Visibility <- "Grzałka"
   TextField "Text field_16" at 472,242 size 69x39; Text 'ppm'
   Circle "Circle_4" at 695,101 size 48x48
      Visibility <- "Pompa_wodna"
   Circle "Circle_5" at 695,243 size 48x48
      Visibility <- "Grzałka"
   Circle "Circle_3" at 695,385 size 48x48
      Visibility <- "Wentylator"
   Circle "Circle_6" at 695,385 size 48x48
      Visibility <- "Wentylator"